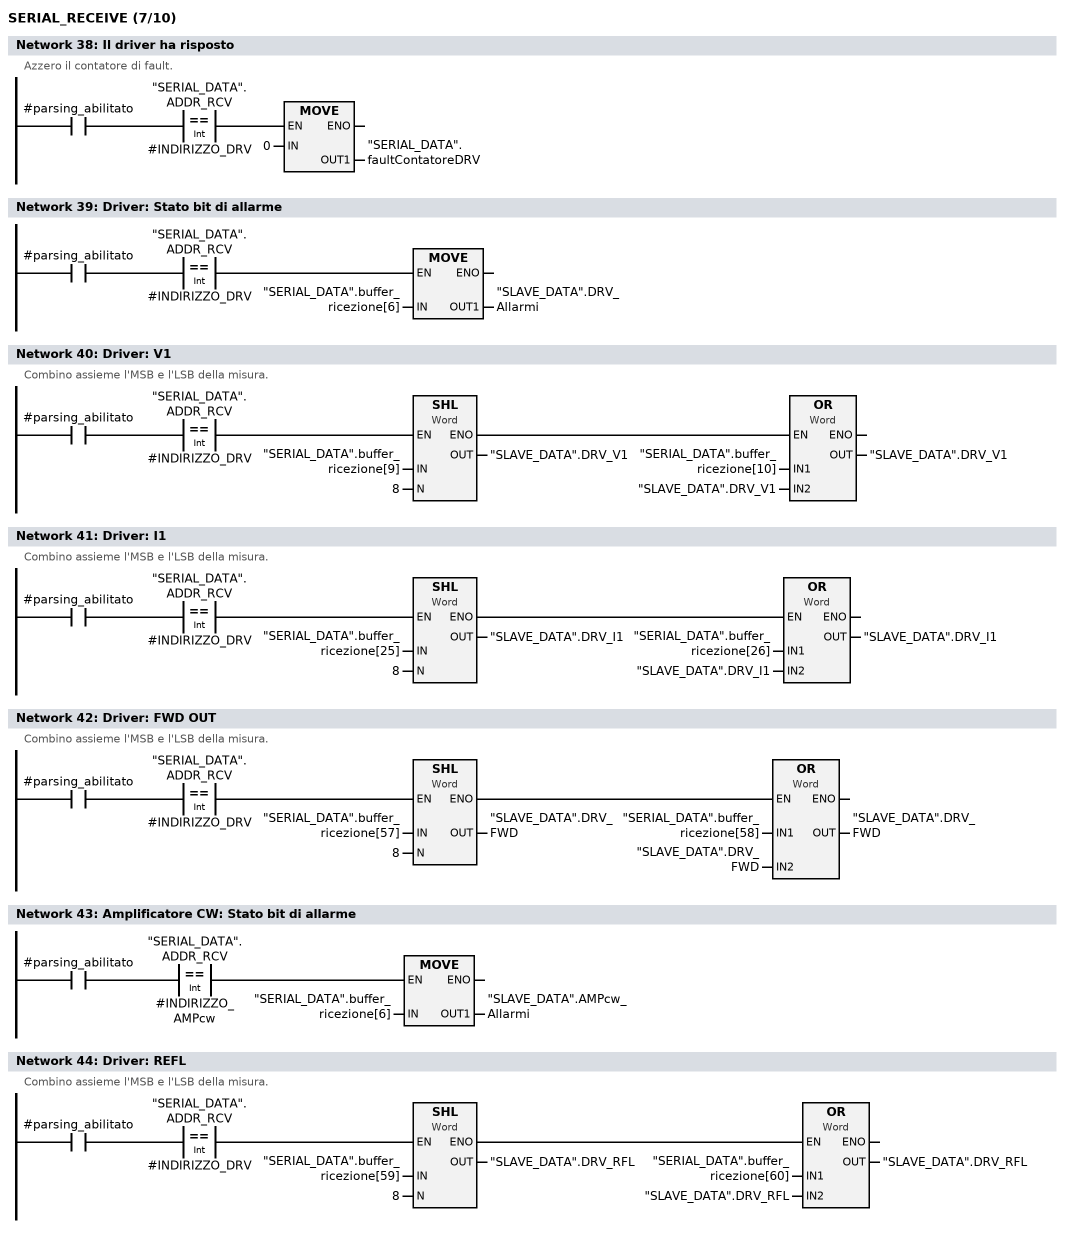
   RUNG wire#powerrail
      Contact( #parsing_abilitato )
      { S7_Templates := "SrcType := Int" } EQ_Contact(in1 := "SERIAL_DATA".ADDR_RCV, in2 := #INDIRIZZO_DRV)
      Move(in := 0, out1 => "SERIAL_DATA".faultContatoreDRV)
   END_RUNG
   // the same network as SCL:
   IF #parsing_abilitato AND ("SERIAL_DATA".ADDR_RCV = #INDIRIZZO_DRV) THEN
       "SERIAL_DATA".faultContatoreDRV := 0;
   END_IF;
END_REGION

REGION Network 39: Driver: Stato bit di allarme
   RUNG wire#powerrail
      Contact( #parsing_abilitato )
      { S7_Templates := "SrcType := Int" } EQ_Contact(in1 := "SERIAL_DATA".ADDR_RCV, in2 := #INDIRIZZO_DRV)
      Move(in := "SERIAL_DATA".buffer_ricezione[6], out1 => "SLAVE_DATA".DRV_Allarmi)
   END_RUNG
   // the same network as SCL:
   IF #parsing_abilitato AND ("SERIAL_DATA".ADDR_RCV = #INDIRIZZO_DRV) THEN
       "SLAVE_DATA".DRV_Allarmi := "SERIAL_DATA".buffer_ricezione[6];
   END_IF;
END_REGION

REGION Network 40: Driver: V1
   // Combino assieme l'MSB e l'LSB della misura.
   // no checked SCL form for this network; see the picture
END_REGION

REGION Network 41: Driver: I1
   // Combino assieme l'MSB e l'LSB della misura.
   // no checked SCL form for this network; see the picture
END_REGION

REGION Network 42: Driver: FWD OUT
   // Combino assieme l'MSB e l'LSB della misura.
   // no checked SCL form for this network; see the picture
END_REGION

REGION Network 43: Amplificatore CW: Stato bit di allarme
   RUNG wire#powerrail
      Contact( #parsing_abilitato )
      { S7_Templates := "SrcType := Int" } EQ_Contact(in1 := "SERIAL_DATA".ADDR_RCV, in2 := #INDIRIZZO_AMPcw)
      Move(in := "SERIAL_DATA".buffer_ricezione[6], out1 => "SLAVE_DATA".AMPcw_Allarmi)
   END_RUNG
   // the same network as SCL:
   IF #parsing_abilitato AND ("SERIAL_DATA".ADDR_RCV = #INDIRIZZO_AMPcw) THEN
       "SLAVE_DATA".AMPcw_Allarmi := "SERIAL_DATA".buffer_ricezione[6];
   END_IF;
END_REGION

REGION Network 44: Driver: REFL
   // Combino assieme l'MSB e l'LSB della misura.
   // no checked SCL form for this network; see the picture
END_REGION

REGION Network 45: Driver: Temperatura Dissipatore
   // Combino assieme l'MSB e l'LSB della misura.
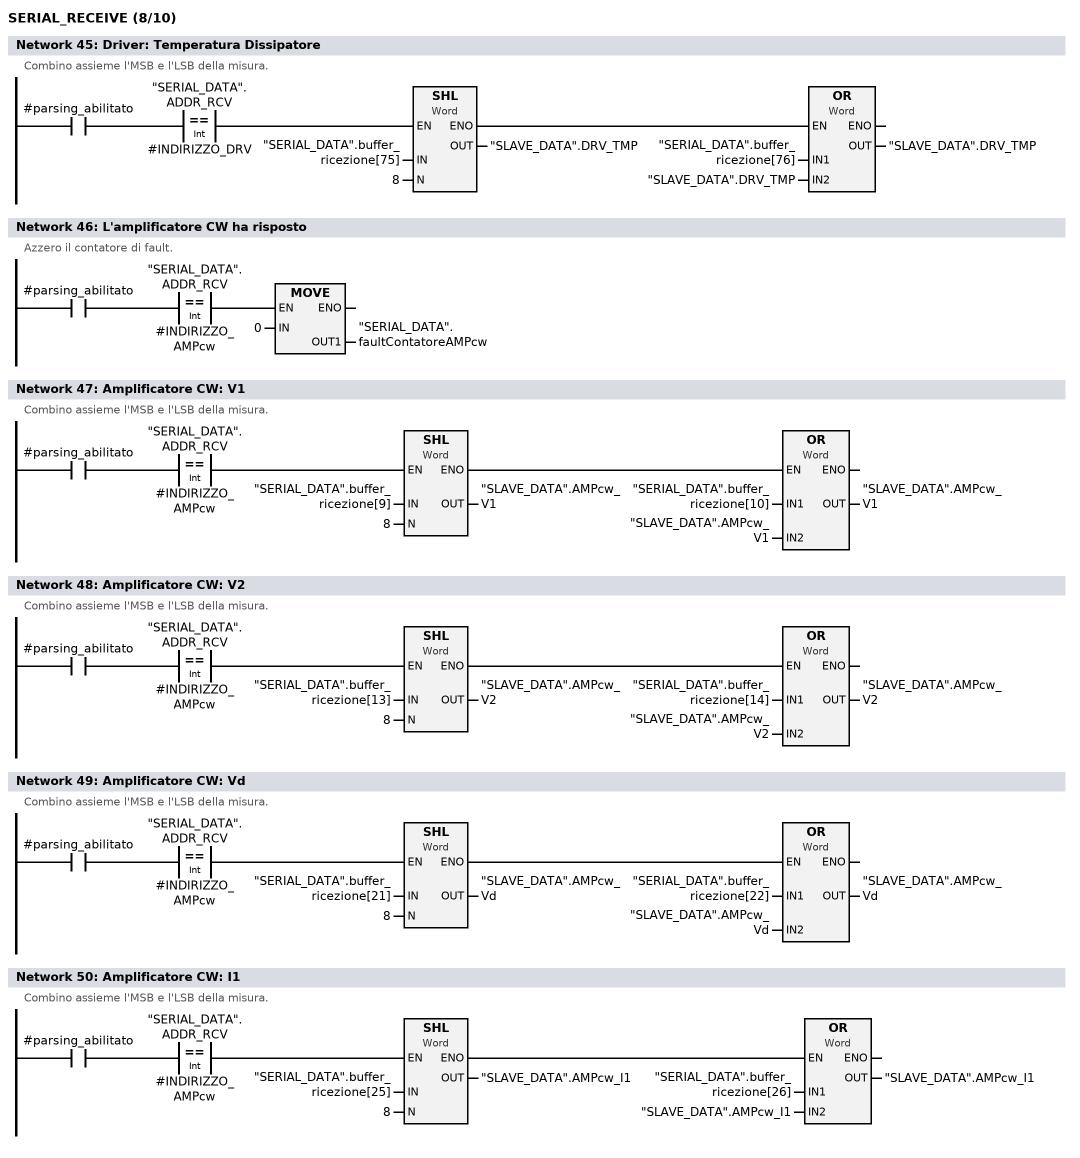
   // no checked SCL form for this network; see the picture
END_REGION

REGION Network 46: L'amplificatore CW ha risposto
   // Azzero il contatore di fault.
   RUNG wire#powerrail
      Contact( #parsing_abilitato )
      { S7_Templates := "SrcType := Int" } EQ_Contact(in1 := "SERIAL_DATA".ADDR_RCV, in2 := #INDIRIZZO_AMPcw)
      Move(in := 0, out1 => "SERIAL_DATA".faultContatoreAMPcw)
   END_RUNG
   // the same network as SCL:
   IF #parsing_abilitato AND ("SERIAL_DATA".ADDR_RCV = #INDIRIZZO_AMPcw) THEN
       "SERIAL_DATA".faultContatoreAMPcw := 0;
   END_IF;
END_REGION

REGION Network 47: Amplificatore CW: V1
   // Combino assieme l'MSB e l'LSB della misura.
   // no checked SCL form for this network; see the picture
END_REGION

REGION Network 48: Amplificatore CW: V2
   // Combino assieme l'MSB e l'LSB della misura.
   // no checked SCL form for this network; see the picture
END_REGION

REGION Network 49: Amplificatore CW: Vd
   // Combino assieme l'MSB e l'LSB della misura.
   // no checked SCL form for this network; see the picture
END_REGION

REGION Network 50: Amplificatore CW: I1
   // Combino assieme l'MSB e l'LSB della misura.
   // no checked SCL form for this network; see the picture
END_REGION

REGION Network 51: Amplificatore CW: I2
   // Combino assieme l'MSB e l'LSB della misura.
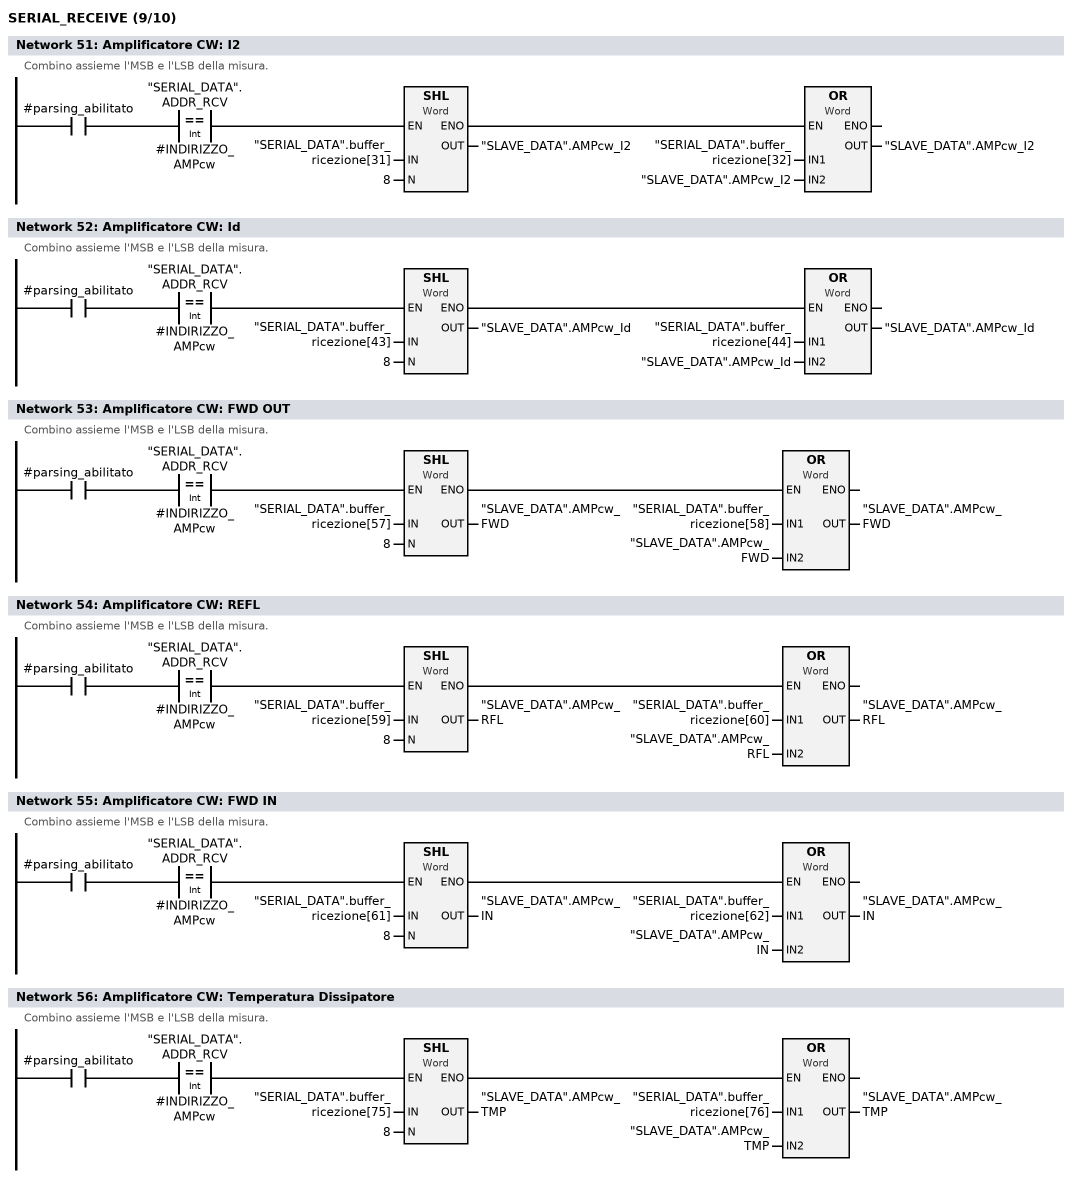
   // no checked SCL form for this network; see the picture
END_REGION

REGION Network 52: Amplificatore CW: Id
   // Combino assieme l'MSB e l'LSB della misura.
   // no checked SCL form for this network; see the picture
END_REGION

REGION Network 53: Amplificatore CW: FWD OUT
   // Combino assieme l'MSB e l'LSB della misura.
   // no checked SCL form for this network; see the picture
END_REGION

REGION Network 54: Amplificatore CW: REFL
   // Combino assieme l'MSB e l'LSB della misura.
   // no checked SCL form for this network; see the picture
END_REGION

REGION Network 55: Amplificatore CW: FWD IN
   // Combino assieme l'MSB e l'LSB della misura.
   // no checked SCL form for this network; see the picture
END_REGION

REGION Network 56: Amplificatore CW: Temperatura Dissipatore
   // Combino assieme l'MSB e l'LSB della misura.
   // no checked SCL form for this network; see the picture
END_REGION

REGION Network 57: Aggiorno l'indirizzo del prossimo slave che deve rispondere
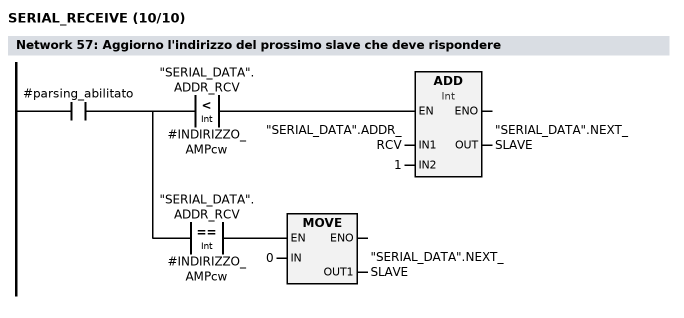
   RUNG wire#powerrail
      Contact( #parsing_abilitato )
      wire#w1
      { S7_Templates := "SrcType := Int" } LT_Contact(in1 := "SERIAL_DATA".ADDR_RCV, in2 := #INDIRIZZO_AMPcw)
      { S7_Templates := "SrcType := Int" } Add(in1 := "SERIAL_DATA".ADDR_RCV, in2 := 1, out => "SERIAL_DATA".NEXT_SLAVE)
   END_RUNG
   RUNG wire#w1
      { S7_Templates := "SrcType := Int" } EQ_Contact(in1 := "SERIAL_DATA".ADDR_RCV, in2 := #INDIRIZZO_AMPcw)
      Move(in := 0, out1 => "SERIAL_DATA".NEXT_SLAVE)
   END_RUNG
   // the same network as SCL:
   IF #parsing_abilitato AND ("SERIAL_DATA".ADDR_RCV < #INDIRIZZO_AMPcw) THEN
       "SERIAL_DATA".NEXT_SLAVE := "SERIAL_DATA".ADDR_RCV + 1;
   END_IF;
   IF #parsing_abilitato AND ("SERIAL_DATA".ADDR_RCV = #INDIRIZZO_AMPcw) THEN
       "SERIAL_DATA".NEXT_SLAVE := 0;
   END_IF;
END_REGION
END_FUNCTION

FUNCTION "ERASE_DATA" : Void   // FC5, LAD
TITLE = ERASE_DATA
{ S7_Optimized_Access := 'FALSE' }
VERSION : 0.1
// Cancella i dati di un blocco se uno slave non risponde in RS485
BEGIN

REGION Network 1: Ricavo l'indirizzo su cui eseguire la cancellazione
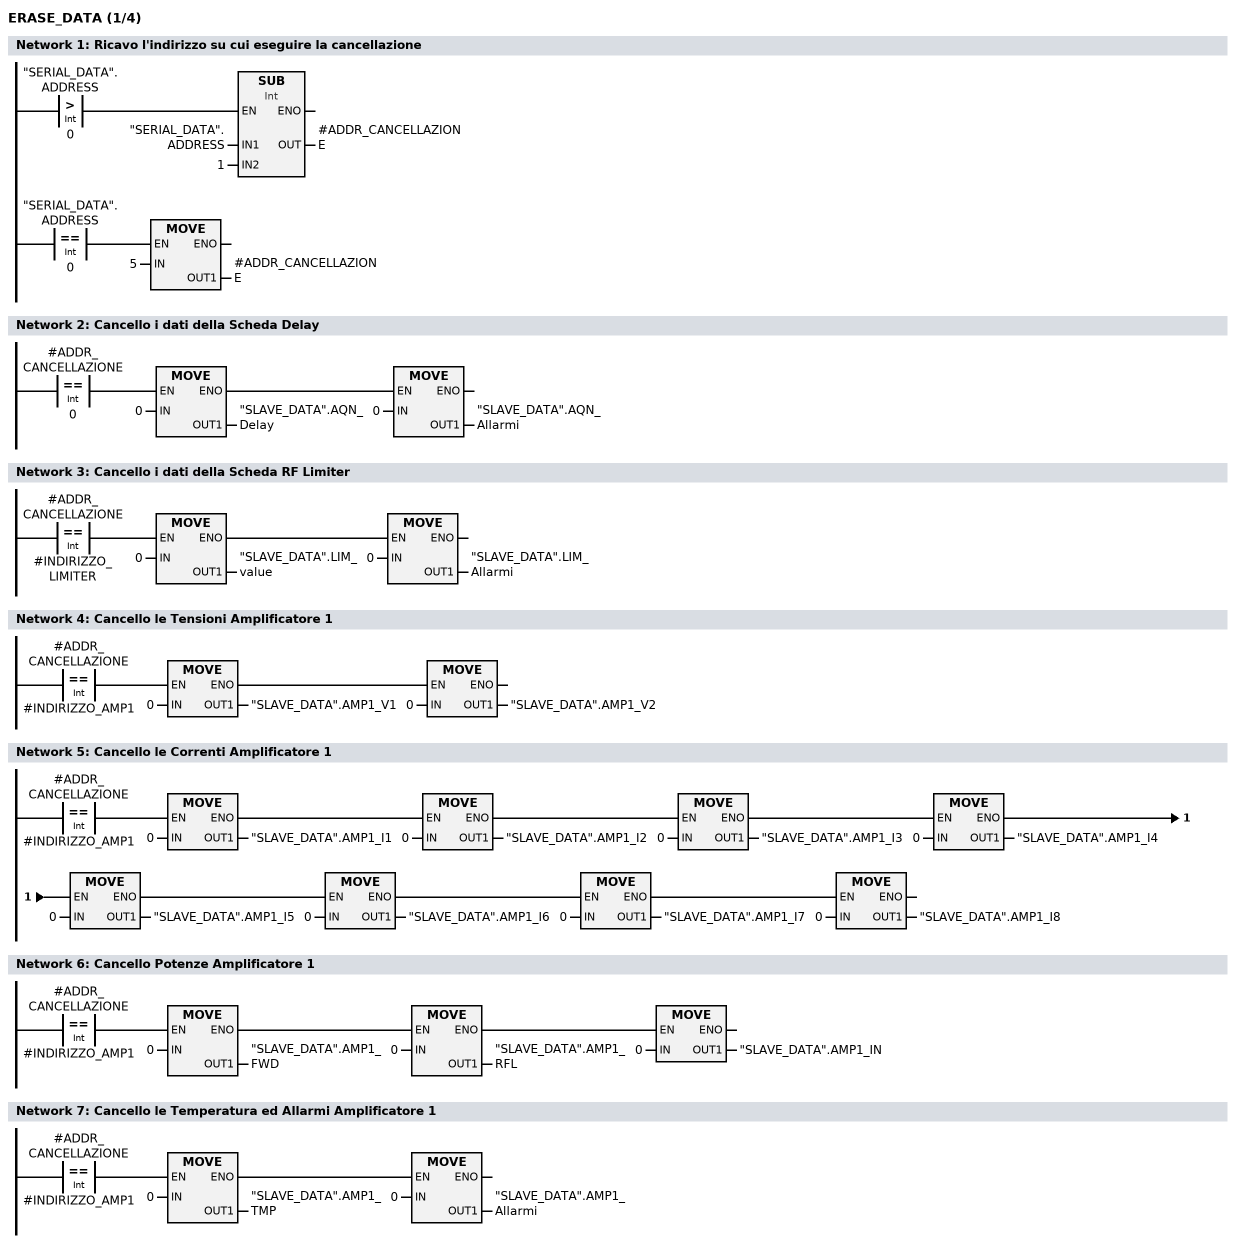
   RUNG wire#powerrail
      { S7_Templates := "SrcType := Int" } GT_Contact(in1 := "SERIAL_DATA".ADDRESS, in2 := 0)
      { S7_Templates := "SrcType := Int" } Sub(in1 := "SERIAL_DATA".ADDRESS, in2 := 1, out => #ADDR_CANCELLAZIONE)
   END_RUNG
   RUNG wire#powerrail
      { S7_Templates := "SrcType := Int" } EQ_Contact(in1 := "SERIAL_DATA".ADDRESS, in2 := 0)
      Move(in := 5, out1 => #ADDR_CANCELLAZIONE)
   END_RUNG
   // the same network as SCL:
   IF "SERIAL_DATA".ADDRESS > 0 THEN #ADDR_CANCELLAZIONE := "SERIAL_DATA".ADDRESS - 1; END_IF;
   IF "SERIAL_DATA".ADDRESS = 0 THEN #ADDR_CANCELLAZIONE := 5; END_IF;
END_REGION

REGION Network 2: Cancello i dati della Scheda Delay
   RUNG wire#powerrail
      { S7_Templates := "SrcType := Int" } EQ_Contact(in1 := #ADDR_CANCELLAZIONE, in2 := 0)
      Move(in := 0, out1 => "SLAVE_DATA".AQN_Delay)
      Move(in := 0, out1 => "SLAVE_DATA".AQN_Allarmi)
   END_RUNG
   // the same network as SCL:
   IF #ADDR_CANCELLAZIONE = 0 THEN
       "SLAVE_DATA".AQN_Delay := 0;
       "SLAVE_DATA".AQN_Allarmi := 0;
   END_IF;
END_REGION

REGION Network 3: Cancello i dati della Scheda RF Limiter
   RUNG wire#powerrail
      { S7_Templates := "SrcType := Int" } EQ_Contact(in1 := #ADDR_CANCELLAZIONE, in2 := #INDIRIZZO_LIMITER)
      Move(in := 0, out1 => "SLAVE_DATA".LIM_value)
      Move(in := 0, out1 => "SLAVE_DATA".LIM_Allarmi)
   END_RUNG
   // the same network as SCL:
   IF #ADDR_CANCELLAZIONE = #INDIRIZZO_LIMITER THEN
       "SLAVE_DATA".LIM_value := 0;
       "SLAVE_DATA".LIM_Allarmi := 0;
   END_IF;
END_REGION

REGION Network 4: Cancello le Tensioni Amplificatore 1
   RUNG wire#powerrail
      { S7_Templates := "SrcType := Int" } EQ_Contact(in1 := #ADDR_CANCELLAZIONE, in2 := #INDIRIZZO_AMP1)
      Move(in := 0, out1 => "SLAVE_DATA".AMP1_V1)
      Move(in := 0, out1 => "SLAVE_DATA".AMP1_V2)
   END_RUNG
   // the same network as SCL:
   IF #ADDR_CANCELLAZIONE = #INDIRIZZO_AMP1 THEN
       "SLAVE_DATA".AMP1_V1 := 0;
       "SLAVE_DATA".AMP1_V2 := 0;
   END_IF;
END_REGION

REGION Network 5: Cancello le Correnti Amplificatore 1
   RUNG wire#powerrail
      { S7_Templates := "SrcType := Int" } EQ_Contact(in1 := #ADDR_CANCELLAZIONE, in2 := #INDIRIZZO_AMP1)
      Move(in := 0, out1 => "SLAVE_DATA".AMP1_I1)
      Move(in := 0, out1 => "SLAVE_DATA".AMP1_I2)
      Move(in := 0, out1 => "SLAVE_DATA".AMP1_I3)
      Move(in := 0, out1 => "SLAVE_DATA".AMP1_I4)
      Move(in := 0, out1 => "SLAVE_DATA".AMP1_I5)
      Move(in := 0, out1 => "SLAVE_DATA".AMP1_I6)
      Move(in := 0, out1 => "SLAVE_DATA".AMP1_I7)
      Move(in := 0, out1 => "SLAVE_DATA".AMP1_I8)
   END_RUNG
   // the same network as SCL:
   IF #ADDR_CANCELLAZIONE = #INDIRIZZO_AMP1 THEN
       "SLAVE_DATA".AMP1_I1 := 0;
       "SLAVE_DATA".AMP1_I2 := 0;
       "SLAVE_DATA".AMP1_I3 := 0;
       "SLAVE_DATA".AMP1_I4 := 0;
       "SLAVE_DATA".AMP1_I5 := 0;
       "SLAVE_DATA".AMP1_I6 := 0;
       "SLAVE_DATA".AMP1_I7 := 0;
       "SLAVE_DATA".AMP1_I8 := 0;
   END_IF;
END_REGION

REGION Network 6: Cancello Potenze Amplificatore 1
   RUNG wire#powerrail
      { S7_Templates := "SrcType := Int" } EQ_Contact(in1 := #ADDR_CANCELLAZIONE, in2 := #INDIRIZZO_AMP1)
      Move(in := 0, out1 => "SLAVE_DATA".AMP1_FWD)
      Move(in := 0, out1 => "SLAVE_DATA".AMP1_RFL)
      Move(in := 0, out1 => "SLAVE_DATA".AMP1_IN)
   END_RUNG
   // the same network as SCL:
   IF #ADDR_CANCELLAZIONE = #INDIRIZZO_AMP1 THEN
       "SLAVE_DATA".AMP1_FWD := 0;
       "SLAVE_DATA".AMP1_RFL := 0;
       "SLAVE_DATA".AMP1_IN := 0;
   END_IF;
END_REGION

REGION Network 7: Cancello le Temperatura ed Allarmi Amplificatore 1
   RUNG wire#powerrail
      { S7_Templates := "SrcType := Int" } EQ_Contact(in1 := #ADDR_CANCELLAZIONE, in2 := #INDIRIZZO_AMP1)
      Move(in := 0, out1 => "SLAVE_DATA".AMP1_TMP)
      Move(in := 0, out1 => "SLAVE_DATA".AMP1_Allarmi)
   END_RUNG
   // the same network as SCL:
   IF #ADDR_CANCELLAZIONE = #INDIRIZZO_AMP1 THEN
       "SLAVE_DATA".AMP1_TMP := 0;
       "SLAVE_DATA".AMP1_Allarmi := 0;
   END_IF;
END_REGION

REGION Network 8: Incremento contatore fault Amplificatore 1
   // Al terzo fault scatta l'allarme.
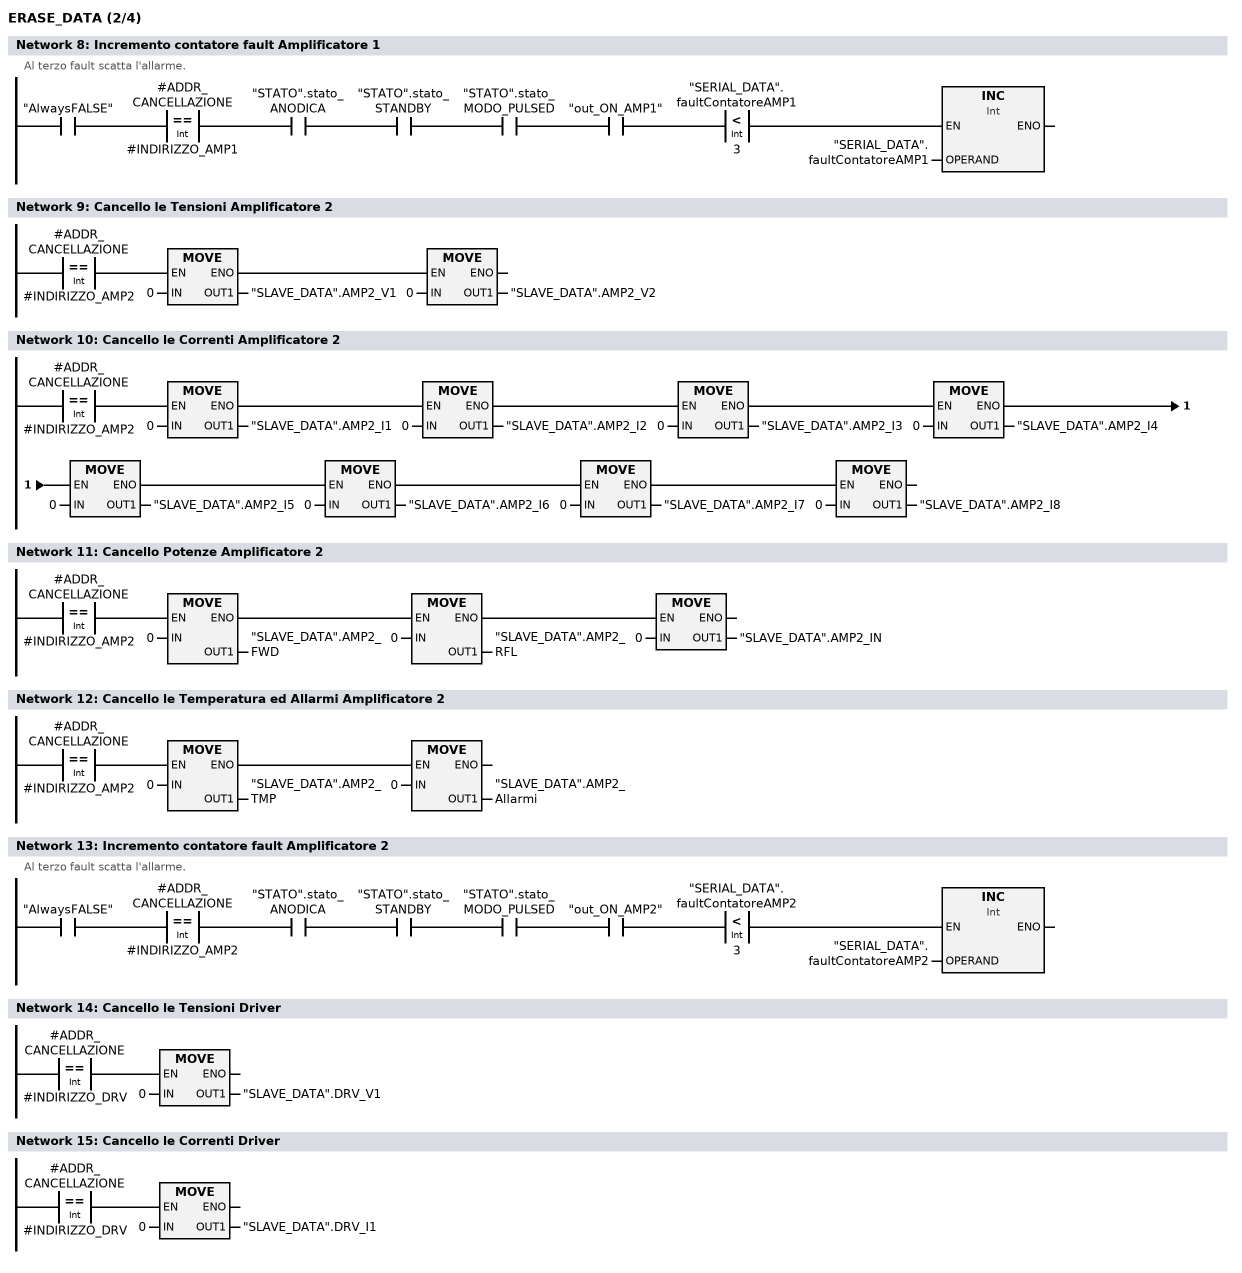
   RUNG wire#powerrail
      Contact( "AlwaysFALSE" )
      { S7_Templates := "SrcType := Int" } EQ_Contact(in1 := #ADDR_CANCELLAZIONE, in2 := #INDIRIZZO_AMP1)
      Contact( "STATO".stato_ANODICA )
      Contact( "STATO".stato_STANDBY )
      Contact( "STATO".stato_MODO_PULSED )
      Contact( "out_ON_AMP1" )
      { S7_Templates := "SrcType := Int" } LT_Contact(in1 := "SERIAL_DATA".faultContatoreAMP1, in2 := 3)
      { S7_Templates := "DestType := Int" } Inc( "SERIAL_DATA".faultContatoreAMP1 )
   END_RUNG
   // the same network as SCL:
   IF "AlwaysFALSE" AND (#ADDR_CANCELLAZIONE = #INDIRIZZO_AMP1) AND "STATO".stato_ANODICA AND "STATO".stato_STANDBY AND "STATO".stato_MODO_PULSED AND "out_ON_AMP1" AND ("SERIAL_DATA".faultContatoreAMP1 < 3) THEN
       "SERIAL_DATA".faultContatoreAMP1 := "SERIAL_DATA".faultContatoreAMP1 + 1;
   END_IF;
END_REGION

REGION Network 9: Cancello le Tensioni Amplificatore 2
   RUNG wire#powerrail
      { S7_Templates := "SrcType := Int" } EQ_Contact(in1 := #ADDR_CANCELLAZIONE, in2 := #INDIRIZZO_AMP2)
      Move(in := 0, out1 => "SLAVE_DATA".AMP2_V1)
      Move(in := 0, out1 => "SLAVE_DATA".AMP2_V2)
   END_RUNG
   // the same network as SCL:
   IF #ADDR_CANCELLAZIONE = #INDIRIZZO_AMP2 THEN
       "SLAVE_DATA".AMP2_V1 := 0;
       "SLAVE_DATA".AMP2_V2 := 0;
   END_IF;
END_REGION

REGION Network 10: Cancello le Correnti Amplificatore 2
   RUNG wire#powerrail
      { S7_Templates := "SrcType := Int" } EQ_Contact(in1 := #ADDR_CANCELLAZIONE, in2 := #INDIRIZZO_AMP2)
      Move(in := 0, out1 => "SLAVE_DATA".AMP2_I1)
      Move(in := 0, out1 => "SLAVE_DATA".AMP2_I2)
      Move(in := 0, out1 => "SLAVE_DATA".AMP2_I3)
      Move(in := 0, out1 => "SLAVE_DATA".AMP2_I4)
      Move(in := 0, out1 => "SLAVE_DATA".AMP2_I5)
      Move(in := 0, out1 => "SLAVE_DATA".AMP2_I6)
      Move(in := 0, out1 => "SLAVE_DATA".AMP2_I7)
      Move(in := 0, out1 => "SLAVE_DATA".AMP2_I8)
   END_RUNG
   // the same network as SCL:
   IF #ADDR_CANCELLAZIONE = #INDIRIZZO_AMP2 THEN
       "SLAVE_DATA".AMP2_I1 := 0;
       "SLAVE_DATA".AMP2_I2 := 0;
       "SLAVE_DATA".AMP2_I3 := 0;
       "SLAVE_DATA".AMP2_I4 := 0;
       "SLAVE_DATA".AMP2_I5 := 0;
       "SLAVE_DATA".AMP2_I6 := 0;
       "SLAVE_DATA".AMP2_I7 := 0;
       "SLAVE_DATA".AMP2_I8 := 0;
   END_IF;
END_REGION

REGION Network 11: Cancello Potenze Amplificatore 2
   RUNG wire#powerrail
      { S7_Templates := "SrcType := Int" } EQ_Contact(in1 := #ADDR_CANCELLAZIONE, in2 := #INDIRIZZO_AMP2)
      Move(in := 0, out1 => "SLAVE_DATA".AMP2_FWD)
      Move(in := 0, out1 => "SLAVE_DATA".AMP2_RFL)
      Move(in := 0, out1 => "SLAVE_DATA".AMP2_IN)
   END_RUNG
   // the same network as SCL:
   IF #ADDR_CANCELLAZIONE = #INDIRIZZO_AMP2 THEN
       "SLAVE_DATA".AMP2_FWD := 0;
       "SLAVE_DATA".AMP2_RFL := 0;
       "SLAVE_DATA".AMP2_IN := 0;
   END_IF;
END_REGION

REGION Network 12: Cancello le Temperatura ed Allarmi Amplificatore 2
   RUNG wire#powerrail
      { S7_Templates := "SrcType := Int" } EQ_Contact(in1 := #ADDR_CANCELLAZIONE, in2 := #INDIRIZZO_AMP2)
      Move(in := 0, out1 => "SLAVE_DATA".AMP2_TMP)
      Move(in := 0, out1 => "SLAVE_DATA".AMP2_Allarmi)
   END_RUNG
   // the same network as SCL:
   IF #ADDR_CANCELLAZIONE = #INDIRIZZO_AMP2 THEN
       "SLAVE_DATA".AMP2_TMP := 0;
       "SLAVE_DATA".AMP2_Allarmi := 0;
   END_IF;
END_REGION

REGION Network 13: Incremento contatore fault Amplificatore 2
   // Al terzo fault scatta l'allarme.
   RUNG wire#powerrail
      Contact( "AlwaysFALSE" )
      { S7_Templates := "SrcType := Int" } EQ_Contact(in1 := #ADDR_CANCELLAZIONE, in2 := #INDIRIZZO_AMP2)
      Contact( "STATO".stato_ANODICA )
      Contact( "STATO".stato_STANDBY )
      Contact( "STATO".stato_MODO_PULSED )
      Contact( "out_ON_AMP2" )
      { S7_Templates := "SrcType := Int" } LT_Contact(in1 := "SERIAL_DATA".faultContatoreAMP2, in2 := 3)
      { S7_Templates := "DestType := Int" } Inc( "SERIAL_DATA".faultContatoreAMP2 )
   END_RUNG
   // the same network as SCL:
   IF "AlwaysFALSE" AND (#ADDR_CANCELLAZIONE = #INDIRIZZO_AMP2) AND "STATO".stato_ANODICA AND "STATO".stato_STANDBY AND "STATO".stato_MODO_PULSED AND "out_ON_AMP2" AND ("SERIAL_DATA".faultContatoreAMP2 < 3) THEN
       "SERIAL_DATA".faultContatoreAMP2 := "SERIAL_DATA".faultContatoreAMP2 + 1;
   END_IF;
END_REGION

REGION Network 14: Cancello le Tensioni Driver
   RUNG wire#powerrail
      { S7_Templates := "SrcType := Int" } EQ_Contact(in1 := #ADDR_CANCELLAZIONE, in2 := #INDIRIZZO_DRV)
      Move(in := 0, out1 => "SLAVE_DATA".DRV_V1)
   END_RUNG
   // the same network as SCL:
   IF #ADDR_CANCELLAZIONE = #INDIRIZZO_DRV THEN "SLAVE_DATA".DRV_V1 := 0; END_IF;
END_REGION

REGION Network 15: Cancello le Correnti Driver
   RUNG wire#powerrail
      { S7_Templates := "SrcType := Int" } EQ_Contact(in1 := #ADDR_CANCELLAZIONE, in2 := #INDIRIZZO_DRV)
      Move(in := 0, out1 => "SLAVE_DATA".DRV_I1)
   END_RUNG
   // the same network as SCL:
   IF #ADDR_CANCELLAZIONE = #INDIRIZZO_DRV THEN "SLAVE_DATA".DRV_I1 := 0; END_IF;
END_REGION

REGION Network 16: Cancello Potenze Driver
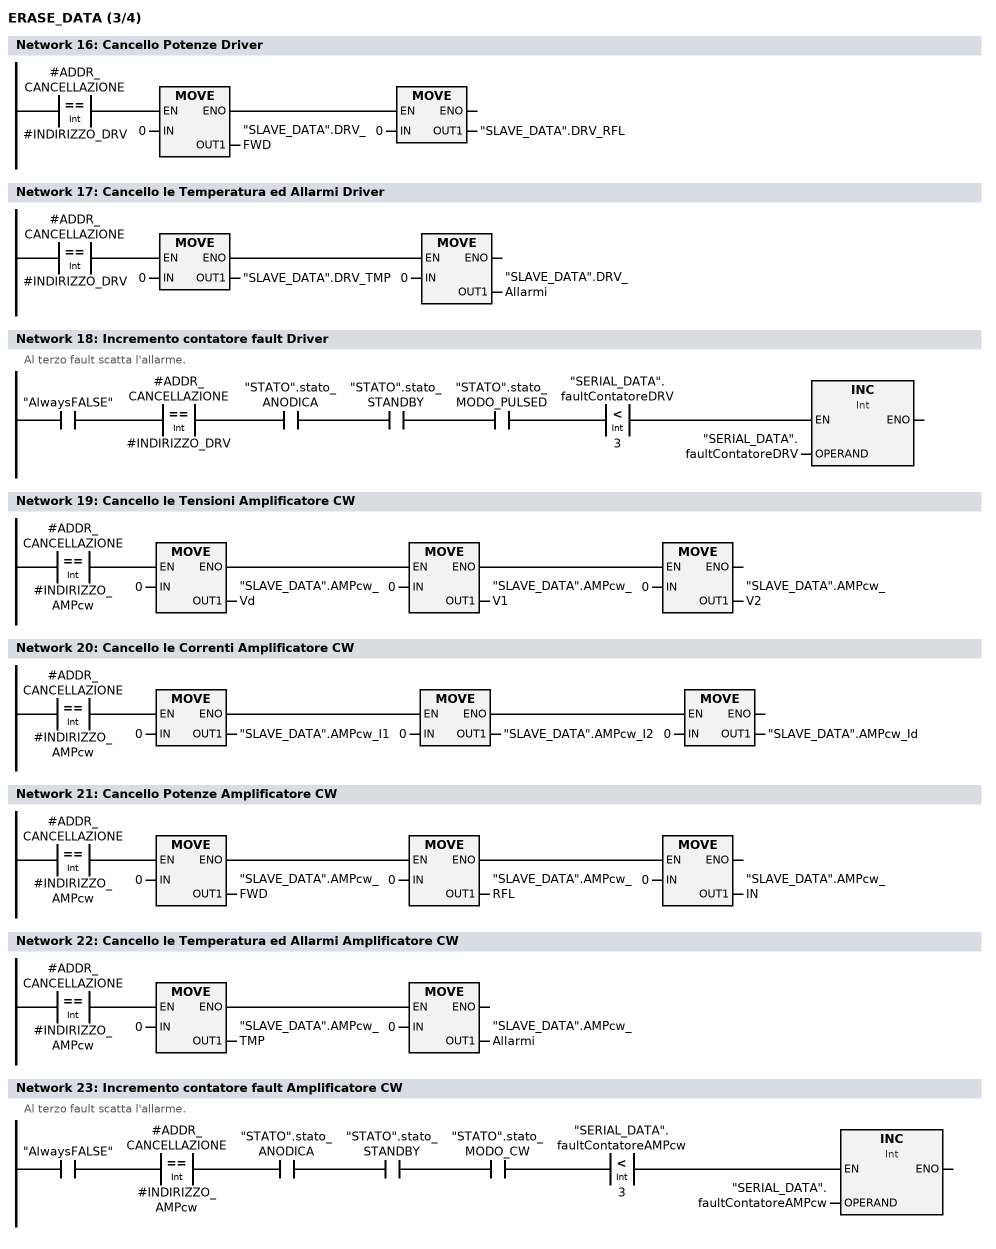
   RUNG wire#powerrail
      { S7_Templates := "SrcType := Int" } EQ_Contact(in1 := #ADDR_CANCELLAZIONE, in2 := #INDIRIZZO_DRV)
      Move(in := 0, out1 => "SLAVE_DATA".DRV_FWD)
      Move(in := 0, out1 => "SLAVE_DATA".DRV_RFL)
   END_RUNG
   // the same network as SCL:
   IF #ADDR_CANCELLAZIONE = #INDIRIZZO_DRV THEN
       "SLAVE_DATA".DRV_FWD := 0;
       "SLAVE_DATA".DRV_RFL := 0;
   END_IF;
END_REGION

REGION Network 17: Cancello le Temperatura ed Allarmi Driver
   RUNG wire#powerrail
      { S7_Templates := "SrcType := Int" } EQ_Contact(in1 := #ADDR_CANCELLAZIONE, in2 := #INDIRIZZO_DRV)
      Move(in := 0, out1 => "SLAVE_DATA".DRV_TMP)
      Move(in := 0, out1 => "SLAVE_DATA".DRV_Allarmi)
   END_RUNG
   // the same network as SCL:
   IF #ADDR_CANCELLAZIONE = #INDIRIZZO_DRV THEN
       "SLAVE_DATA".DRV_TMP := 0;
       "SLAVE_DATA".DRV_Allarmi := 0;
   END_IF;
END_REGION

REGION Network 18: Incremento contatore fault Driver
   // Al terzo fault scatta l'allarme.
   RUNG wire#powerrail
      Contact( "AlwaysFALSE" )
      { S7_Templates := "SrcType := Int" } EQ_Contact(in1 := #ADDR_CANCELLAZIONE, in2 := #INDIRIZZO_DRV)
      Contact( "STATO".stato_ANODICA )
      Contact( "STATO".stato_STANDBY )
      Contact( "STATO".stato_MODO_PULSED )
      { S7_Templates := "SrcType := Int" } LT_Contact(in1 := "SERIAL_DATA".faultContatoreDRV, in2 := 3)
      { S7_Templates := "DestType := Int" } Inc( "SERIAL_DATA".faultContatoreDRV )
   END_RUNG
   // the same network as SCL:
   IF "AlwaysFALSE" AND (#ADDR_CANCELLAZIONE = #INDIRIZZO_DRV) AND "STATO".stato_ANODICA AND "STATO".stato_STANDBY AND "STATO".stato_MODO_PULSED AND ("SERIAL_DATA".faultContatoreDRV < 3) THEN
       "SERIAL_DATA".faultContatoreDRV := "SERIAL_DATA".faultContatoreDRV + 1;
   END_IF;
END_REGION

REGION Network 19: Cancello le Tensioni Amplificatore CW
   RUNG wire#powerrail
      { S7_Templates := "SrcType := Int" } EQ_Contact(in1 := #ADDR_CANCELLAZIONE, in2 := #INDIRIZZO_AMPcw)
      Move(in := 0, out1 => "SLAVE_DATA".AMPcw_Vd)
      Move(in := 0, out1 => "SLAVE_DATA".AMPcw_V1)
      Move(in := 0, out1 => "SLAVE_DATA".AMPcw_V2)
   END_RUNG
   // the same network as SCL:
   IF #ADDR_CANCELLAZIONE = #INDIRIZZO_AMPcw THEN
       "SLAVE_DATA".AMPcw_Vd := 0;
       "SLAVE_DATA".AMPcw_V1 := 0;
       "SLAVE_DATA".AMPcw_V2 := 0;
   END_IF;
END_REGION

REGION Network 20: Cancello le Correnti Amplificatore CW
   RUNG wire#powerrail
      { S7_Templates := "SrcType := Int" } EQ_Contact(in1 := #ADDR_CANCELLAZIONE, in2 := #INDIRIZZO_AMPcw)
      Move(in := 0, out1 => "SLAVE_DATA".AMPcw_I1)
      Move(in := 0, out1 => "SLAVE_DATA".AMPcw_I2)
      Move(in := 0, out1 => "SLAVE_DATA".AMPcw_Id)
   END_RUNG
   // the same network as SCL:
   IF #ADDR_CANCELLAZIONE = #INDIRIZZO_AMPcw THEN
       "SLAVE_DATA".AMPcw_I1 := 0;
       "SLAVE_DATA".AMPcw_I2 := 0;
       "SLAVE_DATA".AMPcw_Id := 0;
   END_IF;
END_REGION

REGION Network 21: Cancello Potenze Amplificatore CW
   RUNG wire#powerrail
      { S7_Templates := "SrcType := Int" } EQ_Contact(in1 := #ADDR_CANCELLAZIONE, in2 := #INDIRIZZO_AMPcw)
      Move(in := 0, out1 => "SLAVE_DATA".AMPcw_FWD)
      Move(in := 0, out1 => "SLAVE_DATA".AMPcw_RFL)
      Move(in := 0, out1 => "SLAVE_DATA".AMPcw_IN)
   END_RUNG
   // the same network as SCL:
   IF #ADDR_CANCELLAZIONE = #INDIRIZZO_AMPcw THEN
       "SLAVE_DATA".AMPcw_FWD := 0;
       "SLAVE_DATA".AMPcw_RFL := 0;
       "SLAVE_DATA".AMPcw_IN := 0;
   END_IF;
END_REGION

REGION Network 22: Cancello le Temperatura ed Allarmi Amplificatore CW
   RUNG wire#powerrail
      { S7_Templates := "SrcType := Int" } EQ_Contact(in1 := #ADDR_CANCELLAZIONE, in2 := #INDIRIZZO_AMPcw)
      Move(in := 0, out1 => "SLAVE_DATA".AMPcw_TMP)
      Move(in := 0, out1 => "SLAVE_DATA".AMPcw_Allarmi)
   END_RUNG
   // the same network as SCL:
   IF #ADDR_CANCELLAZIONE = #INDIRIZZO_AMPcw THEN
       "SLAVE_DATA".AMPcw_TMP := 0;
       "SLAVE_DATA".AMPcw_Allarmi := 0;
   END_IF;
END_REGION

REGION Network 23: Incremento contatore fault Amplificatore CW
   // Al terzo fault scatta l'allarme.
   RUNG wire#powerrail
      Contact( "AlwaysFALSE" )
      { S7_Templates := "SrcType := Int" } EQ_Contact(in1 := #ADDR_CANCELLAZIONE, in2 := #INDIRIZZO_AMPcw)
      Contact( "STATO".stato_ANODICA )
      Contact( "STATO".stato_STANDBY )
      Contact( "STATO".stato_MODO_CW )
      { S7_Templates := "SrcType := Int" } LT_Contact(in1 := "SERIAL_DATA".faultContatoreAMPcw, in2 := 3)
      { S7_Templates := "DestType := Int" } Inc( "SERIAL_DATA".faultContatoreAMPcw )
   END_RUNG
   // the same network as SCL:
   IF "AlwaysFALSE" AND (#ADDR_CANCELLAZIONE = #INDIRIZZO_AMPcw) AND "STATO".stato_ANODICA AND "STATO".stato_STANDBY AND "STATO".stato_MODO_CW AND ("SERIAL_DATA".faultContatoreAMPcw < 3) THEN
       "SERIAL_DATA".faultContatoreAMPcw := "SERIAL_DATA".faultContatoreAMPcw + 1;
   END_IF;
END_REGION

REGION Network 24: Aggiorno l'indirizzo al prossimo slave di cui si attende la risposta
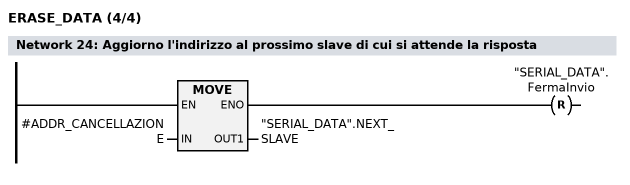
   RUNG wire#powerrail
      Move(in := #ADDR_CANCELLAZIONE, out1 => "SERIAL_DATA".NEXT_SLAVE)
      R_Coil( "SERIAL_DATA".FermaInvio )
   END_RUNG
   // the same network as SCL:
   "SERIAL_DATA".NEXT_SLAVE := #ADDR_CANCELLAZIONE;
   "SERIAL_DATA".FermaInvio := FALSE;
END_REGION
END_FUNCTION

FUNCTION "CALCOLO_LRC_RX" : Void   // FC6, LAD
{ S7_Optimized_Access := 'FALSE' }
VERSION : 0.1
BEGIN

REGION Network 1: Inizializzazione variabili controllo per il calcolo dell'LRC